   //Byte 3
   //Bit                76543210765432107654321076543210         76543210765432107654321076543210
   IF ((#dWordActCycle AND DW#2#00000011000000000000000000000000) = DW#2#00000010000000000000000000000000) THEN
     #tempCount := #tempCount + 1;
   END_IF;
   //Bit                76543210765432107654321076543210         76543210765432107654321076543210
   IF ((#dWordActCycle AND DW#2#00000110000000000000000000000000) = DW#2#00000100000000000000000000000000) THEN
     #tempCount := #tempCount + 1;
   END_IF;
   //Bit                76543210765432107654321076543210         76543210765432107654321076543210
   IF ((#dWordActCycle AND DW#2#00001100000000000000000000000000) = DW#2#00001000000000000000000000000000) THEN
     #tempCount := #tempCount + 1;
   END_IF;
   //Bit                76543210765432107654321076543210         76543210765432107654321076543210
   IF ((#dWordActCycle AND DW#2#00011000000000000000000000000000) = DW#2#00010000000000000000000000000000) THEN
     #tempCount := #tempCount + 1;
   END_IF;
   //Bit                76543210765432107654321076543210         76543210765432107654321076543210
   IF ((#dWordActCycle AND DW#2#00110000000000000000000000000000) = DW#2#00100000000000000000000000000000) THEN
     #tempCount := #tempCount + 1;
   END_IF;
   //Bit                76543210765432107654321076543210         76543210765432107654321076543210
   IF ((#dWordActCycle AND DW#2#01100000000000000000000000000000) = DW#2#01000000000000000000000000000000) THEN
     #tempCount := #tempCount + 1;
   END_IF;
   //Bit                76543210765432107654321076543210         76543210765432107654321076543210
   IF ((#dWordActCycle AND DW#2#11000000000000000000000000000000) = DW#2#10000000000000000000000000000000) THEN
     #tempCount := #tempCount + 1;
   END_IF;
   //Bit                 76543210765432107654321076543210         76543210765432107654321076543210
   IF (((#dWordActCycle AND DW#2#10000000000000000000000000000000) = DW#2#00000000000000000000000000000000)
     AND ((#statDWordPrevCycle AND DW#2#00000000000000000000000000000001) = DW#2#00000000000000000000000000000001))
   THEN
     #tempCount := #tempCount + 1;
   END_IF;

   // Copy DWord actual cycle to DWord previous cycle
   #statDWordPrevCycle := #dWordActCycle;

   //Output
   #countFalInDWord := #tempCount;
END_FUNCTION_BLOCK

FUNCTION_BLOCK "LGF_CountRisInDWordFB"   // FB10004, SCL
{ S7_Optimized_Access := 'TRUE' }
VERSION : 0.1
   VAR_INPUT
      dWordActCycle : DWord;   // Double word in which the rising edges are counted
   END_VAR
   VAR_OUTPUT
      countRisInDWord : Int;   // Number of rising edges in the double word
   END_VAR
   VAR
      statDWordPrevCycle : DWord;   // Double word from the previous cycle
   END_VAR
   VAR_TEMP
      tempCount : Int;
   END_VAR
BEGIN
   //=============================================================================
   // SIEMENS AG
   // (c)Copyright 2017
   //-----------------------------------------------------------------------------
   // Library:       LGF (Library General Functions)
   // Tested with:   CPU1212C DC/DC/DC FW:V4.2
   // Engineering:   TIA Portal V14 Update 1
   // Restrictions:  -
   // Requirements:  PLC (S7-1200 / S7-1500)
   // Functionality: Detects rising edges in variables of type DWORD
   //-----------------------------------------------------------------------------
   // Change log table:
   // Version  Date        In charge / Changes applied
   // 01.00.00 16.01.2019  Siemens Industry Online Support
   //                      First released version
   //=============================================================================

   // Initialization
   #tempCount := 0;

   //Byte 0
   //Bit                76543210765432107654321076543210         76543210765432107654321076543210
   IF ((#dWordActCycle AND DW#2#00000000000000000000000000000011) = DW#2#00000000000000000000000000000001) THEN
     #tempCount := #tempCount + 1;
   END_IF;
   //Bit                76543210765432107654321076543210         76543210765432107654321076543210
   IF ((#dWordActCycle AND DW#2#00000000000000000000000000000110) = DW#2#00000000000000000000000000000010) THEN
     #tempCount := #tempCount + 1;
   END_IF;
   //Bit                76543210765432107654321076543210         76543210765432107654321076543210
   IF ((#dWordActCycle AND DW#2#00000000000000000000000000001100) = DW#2#00000000000000000000000000000100) THEN
     #tempCount := #tempCount + 1;
   END_IF;
   //Bit                76543210765432107654321076543210         76543210765432107654321076543210
   IF ((#dWordActCycle AND DW#2#00000000000000000000000000011000) = DW#2#00000000000000000000000000001000) THEN
     #tempCount := #tempCount + 1;
   END_IF;
   //Bit                76543210765432107654321076543210         76543210765432107654321076543210
   IF ((#dWordActCycle AND DW#2#00000000000000000000000000110000) = DW#2#00000000000000000000000000010000) THEN
     #tempCount := #tempCount + 1;
   END_IF;
   //Bit                76543210765432107654321076543210         76543210765432107654321076543210
   IF ((#dWordActCycle AND DW#2#00000000000000000000000001100000) = DW#2#00000000000000000000000000100000) THEN
     #tempCount := #tempCount + 1;
   END_IF;
   //Bit                76543210765432107654321076543210         76543210765432107654321076543210
   IF ((#dWordActCycle AND DW#2#00000000000000000000000011000000) = DW#2#00000000000000000000000001000000) THEN
     #tempCount := #tempCount + 1;
   END_IF;
   //Bit                76543210765432107654321076543210         76543210765432107654321076543210
   IF ((#dWordActCycle AND DW#2#00000000000000000000000110000000) = DW#2#00000000000000000000000010000000) THEN
     #tempCount := #tempCount + 1;
   END_IF;

   //Byte 1
   //Bit                76543210765432107654321076543210         76543210765432107654321076543210
   IF ((#dWordActCycle AND DW#2#00000000000000000000001100000000) = DW#2#00000000000000000000000100000000) THEN
     #tempCount := #tempCount + 1;
   END_IF;
   //Bit                76543210765432107654321076543210         76543210765432107654321076543210
   IF ((#dWordActCycle AND DW#2#00000000000000000000011000000000) = DW#2#00000000000000000000001000000000) THEN
     #tempCount := #tempCount + 1;
   END_IF;
   //Bit                76543210765432107654321076543210         76543210765432107654321076543210
   IF ((#dWordActCycle AND DW#2#00000000000000000000110000000000) = DW#2#00000000000000000000010000000000) THEN
     #tempCount := #tempCount + 1;
   END_IF;
   //Bit                76543210765432107654321076543210         76543210765432107654321076543210
   IF ((#dWordActCycle AND DW#2#00000000000000000001100000000000) = DW#2#00000000000000000000100000000000) THEN
     #tempCount := #tempCount + 1;
   END_IF;
   //Bit                76543210765432107654321076543210         76543210765432107654321076543210
   IF ((#dWordActCycle AND DW#2#00000000000000000011000000000000) = DW#2#00000000000000000001000000000000) THEN
     #tempCount := #tempCount + 1;
   END_IF;
   //Bit                76543210765432107654321076543210         76543210765432107654321076543210
   IF ((#dWordActCycle AND DW#2#00000000000000000110000000000000) = DW#2#00000000000000000010000000000000) THEN
     #tempCount := #tempCount + 1;
   END_IF;
   //Bit                76543210765432107654321076543210         76543210765432107654321076543210
   IF ((#dWordActCycle AND DW#2#00000000000000001100000000000000) = DW#2#00000000000000000100000000000000) THEN
     #tempCount := #tempCount + 1;
   END_IF;
   //Bit                76543210765432107654321076543210         76543210765432107654321076543210
   IF ((#dWordActCycle AND DW#2#00000000000000011000000000000000) = DW#2#00000000000000001000000000000000) THEN
     #tempCount := #tempCount + 1;
   END_IF;

   //Byte 2
   //Bit                76543210765432107654321076543210         76543210765432107654321076543210
   IF ((#dWordActCycle AND DW#2#00000000000000110000000000000000) = DW#2#00000000000000010000000000000000) THEN
     #tempCount := #tempCount + 1;
   END_IF;
   //Bit                76543210765432107654321076543210         76543210765432107654321076543210
   IF ((#dWordActCycle AND DW#2#00000000000001100000000000000000) = DW#2#00000000000000100000000000000000) THEN
     #tempCount := #tempCount + 1;
   END_IF;
   //Bit                76543210765432107654321076543210         76543210765432107654321076543210
   IF ((#dWordActCycle AND DW#2#00000000000011000000000000000000) = DW#2#00000000000001000000000000000000) THEN
     #tempCount := #tempCount + 1;
   END_IF;
   //Bit                76543210765432107654321076543210         76543210765432107654321076543210
   IF ((#dWordActCycle AND DW#2#00000000000110000000000000000000) = DW#2#00000000000010000000000000000000) THEN
     #tempCount := #tempCount + 1;
   END_IF;
   //Bit                76543210765432107654321076543210         76543210765432107654321076543210
   IF ((#dWordActCycle AND DW#2#00000000001100000000000000000000) = DW#2#00000000000100000000000000000000) THEN
     #tempCount := #tempCount + 1;
   END_IF;
   //Bit                76543210765432107654321076543210         76543210765432107654321076543210
   IF ((#dWordActCycle AND DW#2#00000000011000000000000000000000) = DW#2#00000000001000000000000000000000) THEN
     #tempCount := #tempCount + 1;
   END_IF;
   //Bit                76543210765432107654321076543210         76543210765432107654321076543210
   IF ((#dWordActCycle AND DW#2#00000000110000000000000000000000) = DW#2#00000000010000000000000000000000) THEN
     #tempCount := #tempCount + 1;
   END_IF;
   //Bit                76543210765432107654321076543210         76543210765432107654321076543210
   IF ((#dWordActCycle AND DW#2#00000001100000000000000000000000) = DW#2#00000000100000000000000000000000) THEN
     #tempCount := #tempCount + 1;
   END_IF;

   //Byte 3
   //Bit                76543210765432107654321076543210         76543210765432107654321076543210
   IF ((#dWordActCycle AND DW#2#00000011000000000000000000000000) = DW#2#00000001000000000000000000000000) THEN
     #tempCount := #tempCount + 1;
   END_IF;
   //Bit                76543210765432107654321076543210         76543210765432107654321076543210
   IF ((#dWordActCycle AND DW#2#00000110000000000000000000000000) = DW#2#00000010000000000000000000000000) THEN
     #tempCount := #tempCount + 1;
   END_IF;
   //Bit                76543210765432107654321076543210         76543210765432107654321076543210
   IF ((#dWordActCycle AND DW#2#00001100000000000000000000000000) = DW#2#00000100000000000000000000000000) THEN
     #tempCount := #tempCount + 1;
   END_IF;
   //Bit                76543210765432107654321076543210         76543210765432107654321076543210
   IF ((#dWordActCycle AND DW#2#00011000000000000000000000000000) = DW#2#00001000000000000000000000000000) THEN
     #tempCount := #tempCount + 1;
   END_IF;
   //Bit                76543210765432107654321076543210         76543210765432107654321076543210
   IF ((#dWordActCycle AND DW#2#00110000000000000000000000000000) = DW#2#00010000000000000000000000000000) THEN
     #tempCount := #tempCount + 1;
   END_IF;
   //Bit                76543210765432107654321076543210         76543210765432107654321076543210
   IF ((#dWordActCycle AND DW#2#01100000000000000000000000000000) = DW#2#00100000000000000000000000000000) THEN
     #tempCount := #tempCount + 1;
   END_IF;
   //Bit                76543210765432107654321076543210         76543210765432107654321076543210
   IF ((#dWordActCycle AND DW#2#11000000000000000000000000000000) = DW#2#01000000000000000000000000000000) THEN
     #tempCount := #tempCount + 1;
   END_IF;
   //Bit                 76543210765432107654321076543210         76543210765432107654321076543210
   IF (((#dWordActCycle AND DW#2#10000000000000000000000000000000) = DW#2#10000000000000000000000000000000)
     AND ((#statDWordPrevCycle AND DW#2#00000000000000000000000000000001) = DW#2#00000000000000000000000000000000))
   THEN
     #tempCount := #tempCount + 1;
   END_IF;

   // Copy DWord actual cycle to DWord previous cycle
   #statDWordPrevCycle := #dWordActCycle;

   //Output
   #countRisInDWord := #tempCount;
END_FUNCTION_BLOCK

// folder: Phisical_functions/LGF/3 Comperator operations

FUNCTION "LGF_CompareVariant" : Bool   // FC10005, SCL
{ S7_Optimized_Access := 'FALSE' }
   VAR_OUTPUT
      error : Bool;
      statusID : UInt;
      status : Word;
   END_VAR
   VAR_IN_OUT
      variable1 : Variant;   // First variable
      variable2 : Variant;   // Second variable
   END_VAR
   VAR_TEMP
      tempVariable1Size : DInt;
      tempVariable2Size : DInt;
      tempCounter : DInt;
      tempVariable1ToBytes : Array[1..#MAX_LENGTH] of Byte;
      tempVariable2ToBytes : Array[1..#MAX_LENGTH] of Byte;
      tempSerializeRet : Int;   // Errorcode. Negative if function fails
   END_VAR
   // Ret_Val : TRUE: equal; FALSE: not equal;
   VAR CONSTANT
      NO_ERROR : Word := 16#0000;
      NO_CURRENT_JOBS : Word := 16#7000;
      ERROR_IN_THIS_BLOCK : UInt := 1;
      ERROR_SERIALIZE : UInt := 2;
      MAX_LENGTH : Int := 200;   // Max. length of PLC datatype in Bytes
   END_VAR
BEGIN
   //=============================================================================
   // SIEMENS AG
   // (c)Copyright 2017
   //-----------------------------------------------------------------------------
   // Library:       LGF (Library General Functions)
   // Tested with:   CPU1212C DC/DC/DC FW:V4.2
   // Engineering:   TIA Portal V14 Update 1
   // Restrictions:  -
   // Requirements:  PLC (S7-1200 / S7-1500)
   // Functionality: Compare the datatypes and values up to a max lengh of 200 Bytes
   //                of the connected variables.
   //                If at least one value of an element is not identical -->
   //                set function result = false
   //-----------------------------------------------------------------------------
   // Change log table:
   // Version Date         In charge / Changes applied
   // 01.00.00 03.09.2015  Siemens Industry Online Support
   //                      First released version
   // 01.00.01 11.02.2015  Siemens Industry Online Support
   //                      Bug fix
   // 01.00.02 02.01.2017  Siemens Industry Online Support
   //                      Upgrade: TIA V14 Update 1
   // 01.00.03 17.08.2018  Siemens Industry Online Support
   //                      Upgrade: TIA V15 Update 2
   // 01.00.04 23.11.2018  Siemens Industry Online Support
   //                      Upgrade: TIA V15.1
   //=============================================================================

   // Set "No current job" #status
   #error := false;
   #statusID := #ERROR_IN_THIS_BLOCK;
   #status := #NO_CURRENT_JOBS;

   // Initialisation of function result
   #LGF_CompareVariant := false;

   // Check if the datatypes of the connected tags are identical
   IF TypeOf(#variable1) = TypeOf(#variable2)
   THEN
     #tempVariable1Size := 0;
     #tempSerializeRet := Serialize(SRC_VARIABLE := #variable1, // convert variable Wert1 to array of byte
                                    DEST_ARRAY => #tempVariable1ToBytes,
                                    POS := #tempVariable1Size);

   // Check return value of SERIALIZE
   IF #tempSerializeRet <> 0
     THEN
       #error := true;
       #statusID := #ERROR_SERIALIZE;
       #status := INT_TO_WORD(#tempSerializeRet);
       RETURN; // Finish function if conversion fails

     ELSE
       #tempVariable2Size := 0;
       // Convert variable Wert2 to array of byte
       #tempSerializeRet := Serialize(SRC_VARIABLE := #variable2,
                                      DEST_ARRAY => #tempVariable2ToBytes,
                                      POS := #tempVariable2Size);

       // Check return value of SERIALIZE
       IF #tempSerializeRet <> 0
       THEN
         #error := true;
         #statusID := #ERROR_SERIALIZE;
         #status := INT_TO_WORD(#tempSerializeRet);
         RETURN; // Finish function if conversion fails
       ELSE

         // Compare size of both variables
         IF #tempVariable1Size = #tempVariable2Size
         THEN
           #tempCounter := 1;

           // Compare values of temp. array elements of bytes
           WHILE #tempCounter <= #tempVariable1Size DO

             // Compare bytes till difference detected
             IF #tempVariable1ToBytes[#tempCounter] = #tempVariable2ToBytes[#tempCounter]    
             THEN
               #tempCounter := #tempCounter + 1; // Or end of array reached
             ELSE
               EXIT;
             END_IF;

           END_WHILE;

           #tempCounter := #tempCounter - 1;
           #LGF_CompareVariant := #tempCounter = #tempVariable1Size; // Assign function result

         END_IF;
       END_IF;
     END_IF;
   END_IF;

   #status := #NO_ERROR;
END_FUNCTION

FUNCTION "LGF_CompareReal" : Bool   // FC10037, SCL
{ S7_Optimized_Access := 'TRUE' }
VERSION : 0.1
   VAR_INPUT
      valueA : Real;   // Number to be compared.
      valueB : Real;   // Number to be compared.
   END_VAR
   VAR_OUTPUT
      error : Bool;   // 0: No error. / 1: Error
      status : Word;   // Error information.
   END_VAR
   // Ret_Val : -
   VAR CONSTANT
      EPSILON : Real := 1.0E-06;   // Accuracy with which the two numbers are considered equal
      MAX_RANGE_REAL : Real := 3.402823E+38;   // Maximum range of a REAL number
      ERROR_OVERFLOW : Word := 16#8601;   // Maximum range of a REAL number exceeded
      NO_ERROR : Word := 16#0000;   // No error.
   END_VAR
BEGIN
   //=============================================================================
   // Siemens AG
   // (c)Copyright 2017
   //-----------------------------------------------------------------------------
   // Library:       LGF (Library General Functions)
   // Tested with:   CPU1212C DC/DC/DC FW:V4.2
   // Engineering:   TIA Portal V14 Upd 1
   // Restrictions:  -
   // Requirements:  PLC (S7-1200 / S7-1500)
   // Functionality: This function checks real numbers for parity
   //-----------------------------------------------------------------------------
   // Change log table:
   // Version  Date        In charge / Changes applied
   // 01.00.00 13.01.2017  Siemens Industry Online Support
   //                      First released version
   // 01.00.01 17.08.2018  Siemens Industry Online Support
   //                      Upgrade: TIA V15 Update 2
   // 01.00.02 23.11.2018  Siemens Industry Online Support
   //                      Upgrade: TIA V15.1
   //-----------------------------------------------------------------------------
   //Status Codes: 16#0000 - no error
   //              16#8601 - |valueA|+|valueB| exceeds the maximum range of REAL
   //=============================================================================

   // Reset outputs
   #error := FALSE;
   #status := #NO_ERROR;

   // Initialisation of function result
   #LGF_CompareReal := FALSE;

   // Check |valueA|+|valueB| does not exceed the maximum range of REAL
   IF (ABS(#valueA) + ABS(#valueB)) > #MAX_RANGE_REAL THEN
       #error := TRUE;
       #status := #ERROR_OVERFLOW;
       RETURN;
   END_IF;

   // Approximation
   #LGF_CompareReal := ABS(#valueA - #valueB) <= (#EPSILON * (ABS(#valueA) + ABS(#valueB)));
END_FUNCTION

// folder: Phisical_functions/LGF/4 Math operations

FUNCTION_BLOCK "LGF_MinMaxHistory"   // FB10012, SCL
{ S7_Optimized_Access := 'TRUE' }
   VAR_INPUT
      variable : LReal;
      reset : Bool;
   END_VAR
   VAR_OUTPUT
      minValue : LReal := 1.7976931348623157e+308;
      maxValue : LReal := -1.7976931348623157e+308;
   END_VAR
   VAR
      statMinValue : LReal := 1.7976931348623157e+308;
      statMaxValue : LReal := -1.7976931348623157e+308;
   END_VAR
   VAR CONSTANT
      LREAL_MAX : LReal := 1.7976931348623157e+308;
      LREAL_MIN : LReal := -1.7976931348623157e+308;
   END_VAR
BEGIN
   //=============================================================================
   // SIEMENS AG
   // (c)Copyright 2017
   //-----------------------------------------------------------------------------
   // Library:       LGF (Library General Functions)
   // Tested with:   CPU1212C DC/DC/DC FW:V4.2
   // Engineering:   TIA Portal V14 Update 1
   // Restrictions:  -
   // Requirements:  PLC (S7-1200 / S7-1500)
   // Functionality: This function block saves the minimum and maximum value,
   //                since the start of the block.
   //-----------------------------------------------------------------------------
   // Change log table:
   // Version  Date        In charge / Changes applied
   // 01.00.00 19.08.2015  Siemens Industry Online Support
   //                      First released version
   // 01.00.01 02.01.2017  Siemens Industry Online Support
   //                      Upgrade: TIA Portal V14 Update 1
   //                      Code optimization
   // 01.00.02 17.08.2018  Siemens Industry Online Support
   //                      Upgrade: TIA V15 Update 2
   // 01.00.03 23.11.2018  Siemens Industry Online Support
   //                      Upgrade: TIA V15.1
   //=============================================================================

   // Save min value
   IF (#variable < #statMinValue) THEN
     #statMinValue := #variable;
   END_IF;

   // Save max value
   IF (#variable > #statMaxValue ) THEN
     #statMaxValue := #variable;
   END_IF;

   // If reset is TRUE, min and max value are set to 0
   IF (#reset = TRUE)  THEN
     #statMinValue := #LREAL_MAX;
     #statMaxValue := #LREAL_MIN;
   ELSE
     ;
   END_IF;

   // Ouptput of min and max value
   #minValue := #statMinValue;
   #maxValue := #statMaxValue;
END_FUNCTION_BLOCK

FUNCTION_BLOCK "LGF_Integration"   // FB10043, SCL
{ S7_Optimized_Access := 'TRUE' }
VERSION : 0.1
   VAR_INPUT
      value : Real;   // -
      enable : Bool;   // -
      reset : Bool;   // -
   END_VAR
   VAR_OUTPUT
      integral : Real;   // -
      error : Bool;   // -
      statusID : UInt;   // -
      status : Word;   // Status information / -
   END_VAR
   VAR
      statSysTime : DTL;   // -
      statLastTime : DTL;   // -
      statOldValue : Real;   // -
      statIntegral : Real;   // -
      tempValue : Real;   // -
      tempDeltaTimeT : Time;   // -
      tempDeltaTimeDInt : DInt;   // -
      tempDeltaTimeReal : Real;   // -
      tempRetval : Int;   // -
   END_VAR
   VAR CONSTANT
      ZERO : Real := 0.0;
      NO_ERROR : Word := 16#0000;   // -
      NO_CURRENT_JOBS : Word := 16#7000;   // -
      ERROR_IN_THIS_BLOCK : UInt := 1;   // error in this block
      ERROR_RD_SYS_T : UInt := 2;   // error in RD_SYS_T
   END_VAR
BEGIN
   //=============================================================================
   // SIEMENS AG
   // (c)Copyright 2017
   //-----------------------------------------------------------------------------
   // Library:       LGF (Library General Functions)
   // Tested with:   CPU1212C DC/DC/DC FW:V4.2
   // Engineering:   TIA Portal V14 Upd 1
   // Restrictions:  -
   // Requirements:  PLC (S7-1200 / S7-1500)
   // Functionality: The input value will be integrated.
   //                
   //-----------------------------------------------------------------------------
   // Change log table:
   // Version  Date        In charge Changes applied
   // 01.00.00 17.02.2017  Siemens Industry Online Support
   //                      First released version
   // 01.00.01 17.08.2018  Siemens Industry Online Support
   //                      Upgrade: TIA V15 Update 2
   // 01.00.02 23.11.2018  Siemens Industry Online Support
   //                      Upgrade: TIA V15.1
   //-----------------------------------------------------------------------------
   //=============================================================================

   // Initialization
   #error := FALSE;
   #statusID := #NO_ERROR;
   #status := #NO_CURRENT_JOBS;

   // Reset 
   IF #reset = true THEN
     #integral := #ZERO;
     #statOldValue := #ZERO;
     #statIntegral := #ZERO;
     RETURN;
   END_IF;

   // Write input value to temp variable
   #tempValue := #value;

   // Read system time
   #tempRetval := RD_SYS_T(OUT => #statSysTime);

   // Error Handling read system time
   IF (#tempRetval > 1) THEN
     #error := TRUE;
     #statusID := #ERROR_RD_SYS_T;
     #status := INT_TO_WORD(#tempRetval);
     RETURN;
   END_IF;

   // Calculate time difference between last and actual time
   #tempDeltaTimeT := #statSysTime - #statLastTime;

   // Convert times difference to REAL
   #tempDeltaTimeDInt := TIME_TO_DINT(#tempDeltaTimeT);
   #tempDeltaTimeReal := DINT_TO_REAL(#tempDeltaTimeDInt);

   // Convert in seconds
   #tempDeltaTimeReal := #tempDeltaTimeReal / 1000.0;

   // Write actual to last time
   #statLastTime := #statSysTime;

   IF NOT #enable = true THEN
     #statOldValue := #ZERO;
     RETURN;
   END_IF;

   // Add LastScalIn to ScalIn
   #tempValue := #tempValue + #statOldValue;

   // Save last input
   #statOldValue := #value;

   // Divide in half statScalIn
   #tempValue := #tempValue / 2.0;

   // Multiply with Delta Time
   #tempValue := #tempValue * #tempDeltaTimeReal;

   // Calculate new integral
   #statIntegral := #statIntegral + #tempValue;

   // Write outputs
   #integral := #statIntegral;
   #status := #NO_ERROR;
END_FUNCTION_BLOCK

FUNCTION "LGF_RandomInt" : Int   // FC2, SCL
{ S7_Optimized_Access := 'TRUE' }
   VAR_INPUT
      minValue : Int;   // minimal Value random can reach
      maxValue : Int;   // maximal Value random can reach
   END_VAR
   VAR_OUTPUT
      error : Bool;
      statusID : UInt;
      status : Word;
   END_VAR
   VAR_TEMP
      tempTime : DTL;
      tempTimeStatus : Int;
      tempRandomValue : Int;
      tempNormReal : Real;
   END_VAR
   VAR CONSTANT
      NO_ERROR : Word := 16#0000;
      NO_CURRENT_JOBS : Word := 16#7000;
      MAX_LESS_MIN : Word := 16#8200;
      ERROR_IN_THIS_BLOCK : UInt := 1;
      ERROR_RD_SYS_T : UInt := 2;
      MIN_INT : DInt := -32768;
      MAX_INT : DInt := 32767;
   END_VAR
BEGIN
   //=============================================================================
   // Siemens AG
   // (c)Copyright 2017
   //-----------------------------------------------------------------------------
   // Library:       LGF (Library General Functions)
   // Tested with:   CPU1212C DC/DC/DC FW:V4.2
   // Engineering:   TIA Portal V13 SP1 Upd 4
   // Restrictions:  -
   // Requirements:  PLC (S7-1200 / S7-1500)
   // Functionality: This function generates random numbers in defined limits
   //                (Datatype Int)
   //-----------------------------------------------------------------------------
   // Change log table:
   // Version  Date        In charge / Changes applied
   // 01.00.00 19.08.2015  Siemens Industry Online Support
   //                      First released version
   // 01.00.01 02.01.2017  Siemens Industry Online Support
   //                      Upgrade: TIA Portal V14 Update 1
   // 01.00.02 17.08.2018  Siemens Industry Online Support
   //                      Upgrade: TIA V15 Update 2
   // 01.00.03 23.11.2018  Siemens Industry Online Support
   //                      Upgrade: TIA V15.1
   //-----------------------------------------------------------------------------
   //Status Codes:
   // 16#7000:  No current jobs
   // 16#0000:  Job finished; Note: There is no "Busy"-Status because the block
   //           is finished within a single cycle
   // 16#8200:  maxValue is samller then minValue 
   //=============================================================================

   //Set "No current job" status
   #error := false;
   #statusID := #ERROR_IN_THIS_BLOCK;
   #status := #NO_CURRENT_JOBS;

   //Check if the maximal Value is less than the minimal value
   IF (#minValue > #maxValue) THEN
     #error := true;
     #statusID := #ERROR_IN_THIS_BLOCK;
     #status := #MAX_LESS_MIN;
     #LGF_RandomInt := 0;
     RETURN;
   END_IF;

   //Read system time
   #tempTimeStatus := RD_SYS_T(#tempTime);

   IF (#tempTimeStatus <> 0) THEN
     #error := true;
     #statusID := #ERROR_RD_SYS_T;
     #status := INT_TO_WORD(#tempTimeStatus);
     #LGF_RandomInt := 0;
     RETURN;
   END_IF;

   //Callculate a random-start-value depending on the time
   #tempRandomValue.%B1 := #tempTime.NANOSECOND.%B0;
   #tempRandomValue.%B0 := #tempTime.NANOSECOND.%B1;

   //adapt the calculated random number to the given number span
   #tempNormReal := NORM_X(MIN := #MIN_INT, VALUE := #tempRandomValue, MAX := #MAX_INT);
   #LGF_RandomInt := SCALE_X(MIN := #minValue, VALUE := #tempNormReal, MAX := #maxValue);

   #status := #NO_ERROR;
END_FUNCTION

FUNCTION "LGF_Factorial" : DInt   // FC9, SCL
{ S7_Optimized_Access := 'TRUE' }
VERSION : 0.1
   VAR_INPUT
      n : Int;   // Natural number
   END_VAR
   VAR_OUTPUT
      status : Word;   // Status
      error : Bool;   // Error
   END_VAR
   VAR_TEMP
      tempFactorial : DInt;   // Temp Factorial
      tempIndex : Int;   // Temp index
   END_VAR
   // Ret_Val : Calculated factorial
   VAR CONSTANT
      NO_ERROR : Word := 16#0000;   // Status no error
      NO_CURRENT_JOBS : Word := 16#7000;   // Status no current jobs
      WRONG_VALUE_RANGE : Word := 16#8101;   // Status wrong value range for input value
   END_VAR
BEGIN
   //=============================================================================
   // Siemens AG
   // (c)Copyright 2017
   //-----------------------------------------------------------------------------
   // Library:       LGF (Library General Functions)
   // Tested with:   CPU1212C DC/DC/DC FW:V4.2
   // Engineering:   TIA Portal V14 SP1 Upd 5
   // Restrictions:  -
   // Requirements:  PLC (S7-1200 / S7-1500)
   // Functionality: This program calculates factorial values from 1 to 12.
   //-----------------------------------------------------------------------------
   // Change log table:
   // Version  Date        In charge / Changes applied
   // 01.00.00 03.07.2018  Siemens Industry Online Support
   //                      First released version
   // 01.00.01 17.08.2018  Siemens Industry Online Support
   //                      Upgrade: TIA V15 Update 2
   // 01.00.02 23.11.2018  Siemens Industry Online Support
   //                      Upgrade: TIA V15.1
   //-----------------------------------------------------------------------------
   //Status Codes:
   // 16#0000:  Job finished   // Note: There is no "Busy"-Status because the
   //           block is finished within a single cycle
   // 16#8101:  Outside value range ( factorial until 12 is possible)
   //=============================================================================

   #error := FALSE;
   #status := #NO_CURRENT_JOBS;

   IF (#n < 13)
     AND (#n >= 0)
   THEN
     IF (#n = 0)
     THEN
       #tempFactorial := 1;
     ELSE
       #tempFactorial := 1;
       FOR #tempIndex := 1 TO #n DO
         #tempFactorial := #tempFactorial * #tempIndex;
       END_FOR;
     END_IF;

     #error := FALSE; // No errors
     #status := #NO_ERROR;

   ELSE
     #tempFactorial := 0;
     #error := TRUE;
     #status := #WRONG_VALUE_RANGE;
   END_IF;

   #LGF_Factorial := #tempFactorial;
END_FUNCTION

FUNCTION "LGF_MatrixAddition" : Void   // FC10007, SCL
{ S7_Optimized_Access := 'TRUE' }
   VAR_INPUT
      matrix1 : Array[*, *] of Real;   // first summand
      matrix2 : Array[*, *] of Real;   // second summand
   END_VAR
   VAR_OUTPUT
      matrixResult : Array[*, *] of Real;   // result matrix
      error : Bool;
      statusID : UInt;
      status : Word;
   END_VAR
   VAR_TEMP
      tempMatrix1LowerBound1Dim : DInt;   // -
      tempMatrix1LowerBound2Dim : DInt;   // -
      tempMatrix1UpperBound1Dim : DInt;   // -
      tempMatrix1UpperBound2Dim : DInt;   // -
      tempMatrix2LowerBound1Dim : DInt;   // -
      tempMatrix2LowerBound2Dim : DInt;   // -
      tempMatrix2UpperBound1Dim : DInt;   // -
      tempMatrix2UpperBound2Dim : DInt;   // -
      tempResultMatrixLowerBound1Dim : DInt;   // -
      tempResultMatrixLowerBound2Dim : DInt;   // -
      tempResultMatrixUpperBound1Dim : DInt;   // -
      tempResultMatrixUpperBound2Dim : DInt;   // -
      tempCounterDim1 : Int;   // -
      tempCounterDim2 : Int;   // -
   END_VAR
   VAR CONSTANT
      NO_ERROR : Word := 16#0000;   // No errors.
      ERROR_LOWER_BOUND_NOT_EQUAL : Word := 16#8200;   // Lower bounds of matrices are not equal.
      ERROR_UPPER_BOUND_NOT_EQUAL : Word := 16#8201;   // Upper bounds of matrices are not equal.
      ERROR_IN_THIS_BLOCK : UInt := 1;   // statusID: Error in this block.
   END_VAR
BEGIN
   //=============================================================================
   // SIEMENS AG
   // (c)Copyright 2017
   //-----------------------------------------------------------------------------
   // Library:       LGF (Library General Functions)
   // Tested with:   CPU1212C DC/DC/DC FW:V4.2
   // Engineering:   TIA Portal V14 Update 1
   // Restrictions:  -
   // Requirements:  PLC (S7-1200 / S7-1500)
   // Functionality: This function add up matrices.
   //-----------------------------------------------------------------------------
   // Change log table:
   // Version  Date        In charge / Changes applied
   // 01.00.00 19.08.2015  Siemens Industry Online Support
   //                      First released version
   // 01.00.01 02.01.2017  Siemens Industry Online Support
   //                      Upgrade: TIA Portal V14 Update 1
   // 02.00.00 06.02.2017  Siemens Industry Online Support
   //                      Functionality using Array[*,*]
   // 02.00.01 17.08.2018  Siemens Industry Online Support
   //                      Upgrade: TIA V15 Update 2
   // 02.00.02 23.11.2018  Siemens Industry Online Support
   //                      Upgrade: TIA V15.1
   //=============================================================================

   //Set "No error" status
   #error := false;
   #statusID := #ERROR_IN_THIS_BLOCK;
   #status := #NO_ERROR;

   // Init resultMatrix
   #matrixResult[0, 0] := 0.0;

   //Determine the size of the matrices
   // Lower bound dimension 1
   #tempMatrix1LowerBound1Dim := LOWER_BOUND(ARR := #matrix1, DIM := 1);
   #tempMatrix2LowerBound1Dim := LOWER_BOUND(ARR := #matrix2, DIM := 1);
   #tempResultMatrixLowerBound1Dim := LOWER_BOUND(ARR := #matrixResult, DIM := 1);
   // Lower bound dimension 2
   #tempMatrix1LowerBound2Dim := LOWER_BOUND(ARR := #matrix1, DIM := 2);
   #tempMatrix2LowerBound2Dim := LOWER_BOUND(ARR := #matrix2, DIM := 2);
   #tempResultMatrixLowerBound2Dim := LOWER_BOUND(ARR := #matrixResult, DIM := 2);
   // Upper bound dimension 1
   #tempMatrix1UpperBound1Dim := UPPER_BOUND(ARR := #matrix1, DIM := 1);
   #tempMatrix2UpperBound1Dim := UPPER_BOUND(ARR := #matrix2, DIM := 1);
   #tempResultMatrixUpperBound1Dim := UPPER_BOUND(ARR := #matrixResult, DIM := 1);
   // Upper bound dimension 2
   #tempMatrix1UpperBound2Dim := UPPER_BOUND(ARR := #matrix1, DIM := 2);
   #tempMatrix2UpperBound2Dim := UPPER_BOUND(ARR := #matrix2, DIM := 2);
   #tempResultMatrixUpperBound2Dim := UPPER_BOUND(ARR := #matrixResult, DIM := 2);

   // Check the lower bound of all matrices
   IF (#tempMatrix1LowerBound1Dim <> #tempMatrix2LowerBound1Dim) OR (#tempMatrix1LowerBound1Dim <> #tempResultMatrixLowerBound1Dim) OR
     (#tempMatrix1LowerBound2Dim <> #tempMatrix2LowerBound2Dim) OR (#tempMatrix1LowerBound2Dim <> #tempResultMatrixLowerBound2Dim) THEN
     #error := TRUE;
     #status := #ERROR_LOWER_BOUND_NOT_EQUAL;
     RETURN;
   END_IF;
   // Check the upper bound of all matrices
   IF (#tempMatrix1UpperBound1Dim <> #tempMatrix2UpperBound1Dim) OR (#tempMatrix1UpperBound1Dim <> #tempResultMatrixUpperBound1Dim) OR
     (#tempMatrix1UpperBound2Dim <> #tempMatrix2UpperBound2Dim) OR (#tempMatrix1UpperBound2Dim <> #tempResultMatrixUpperBound2Dim) THEN
     #error := TRUE;
     #status := #ERROR_UPPER_BOUND_NOT_EQUAL;
     RETURN;
   END_IF;

   // Addition of two matrices
   FOR #tempCounterDim1 := #tempMatrix1LowerBound1Dim TO #tempMatrix1UpperBound1Dim DO
     FOR #tempCounterDim2 := #tempMatrix1LowerBound2Dim TO #tempMatrix1UpperBound2Dim DO
       #matrixResult[#tempCounterDim1, #tempCounterDim2] := #matrix1[#tempCounterDim1, #tempCounterDim2] + #matrix2[#tempCounterDim1, #tempCounterDim2];
     END_FOR;
   END_FOR;
END_FUNCTION

FUNCTION "LGF_MatrixInverse" : Void   // FC10008, SCL
{ S7_Optimized_Access := 'TRUE' }
   VAR_INPUT
      matrix : Array[*, *] of Real;   // input matrix
   END_VAR
   VAR_OUTPUT
      matrixResult : Array[*, *] of Real;   // output matrix
      error : Bool;
      statusID : UInt;
      status : Word;
   END_VAR
   VAR_TEMP
      tempCounterDim2 : Int;   // -
      tempCounterDim1 : Int;   // -
      tempMatrixLowerBound1Dim : DInt;   // -
      tempMatrixLowerBound2Dim : DInt;   // -
      tempMatrixUpperBound1Dim : DInt;   // -
      tempMatrixUpperBound2Dim : DInt;   // -
      tempResultMatrixLowerBound1Dim : DInt;   // -
      tempResultMatrixLowerBound2Dim : DInt;   // -
      tempResultMatrixUpperBound1Dim : DInt;   // -
      tempResultMatrixUpperBound2Dim : DInt;   // -
      tempColumns : DInt;   // -
      tempRows : DInt;   // -
      tempK : DInt;   // -
      tempI : DInt;   // -
      tempJ : DInt;   // -
   END_VAR
   VAR CONSTANT
      NO_ERROR : Word := 16#0000;   // No error.
      ERROR_LOWER_BOUND_NOT_EQUAL : Word := 16#8200;   // Lower bounds of matrices are not equal.
      ERROR_UPPER_BOUND_NOT_EQUAL : Word := 16#8201;   // Upper bounds of matrices are not equal.
      ERROR_NOT_SQUARE_MATRIX : Word := 16#8202;   // Input matrix is not a square matrix.
      ERROR_ALGORITHM_NOT_POSSIBLE : Word := 16#8203;   // Algorithm not possible for the input matrix.
      ERROR_IN_THIS_BLOCK : UInt := 1;   // statusID: error in this block.
   END_VAR
BEGIN
   //=============================================================================
   // SIEMENS AG
   // (c)Copyright 2017
   //-----------------------------------------------------------------------------
   // Library:       LGF (Library General Functions)
   // Tested with:   CPU1212C DC/DC/DC FW:V4.2
   // Engineering:   TIA Portal V14 Update 1
   // Restrictions:  -
   // Requirements:  PLC (S7-1200 / S7-1500)
   // Functionality: This function inverses matrices. Inversion of regulary,
   //                quadratic Matrix with the Shipley-Coleman method.
   //-----------------------------------------------------------------------------
   // Change log table:
   // Version  Date        In charge / Changes applied
   // 01.00.00 19.08.2015  Siemens Industry Online Support
   //                      First released version
   // 01.00.01 02.01.2017  Siemens Industry Online Support
   //                      Upgrade: TIA Portal V14 Update 1
   // 02.00.00 06.02.2017  Siemens Industry Online Support
   //                      Functionality using Array[*,*]
   // 02.00.01 17.08.2018  Siemens Industry Online Support
   //                      Upgrade: TIA V15 Update 2
   // 02.00.02 23.11.2018  Siemens Industry Online Support
   //                      Upgrade: TIA V15.1
   //=============================================================================

   //Set "No error" status
   #error := false;
   #statusID := #ERROR_IN_THIS_BLOCK;
   #status := #NO_ERROR;

   // Initialize result matrix
   #matrixResult[0, 0] := 0.0;

   //Determine the size of the matrices
   // Lower bound dimension 1
   #tempMatrixLowerBound1Dim := LOWER_BOUND(ARR := #matrix, DIM := 1);
   #tempResultMatrixLowerBound1Dim := LOWER_BOUND(ARR := #matrixResult, DIM := 1);
   // Lower bound dimension 2
   #tempMatrixLowerBound2Dim := LOWER_BOUND(ARR := #matrix, DIM := 2);
   #tempResultMatrixLowerBound2Dim := LOWER_BOUND(ARR := #matrixResult, DIM := 2);
   // Upper bound dimension 1
   #tempMatrixUpperBound1Dim := UPPER_BOUND(ARR := #matrix, DIM := 1);
   #tempResultMatrixUpperBound1Dim := UPPER_BOUND(ARR := #matrixResult, DIM := 1);
   // Upper bound dimension 2
   #tempMatrixUpperBound2Dim := UPPER_BOUND(ARR := #matrix, DIM := 2);
   #tempResultMatrixUpperBound2Dim := UPPER_BOUND(ARR := #matrixResult, DIM := 2);

   // Count the columns of input matrix
   IF #tempMatrixLowerBound2Dim = 0 THEN
     #tempColumns := #tempMatrixUpperBound2Dim + 1;
   ELSE
     #tempColumns := (#tempMatrixUpperBound2Dim - #tempMatrixLowerBound2Dim) + 1;
   END_IF;
   // Count the rows of input matrix
   IF #tempMatrixLowerBound1Dim = 0 THEN
     #tempRows := #tempMatrixUpperBound1Dim + 1;
   ELSE
     #tempRows := (#tempMatrixUpperBound1Dim - #tempMatrixLowerBound1Dim) + 1;
   END_IF;
   // Check whether input matrix is a square matrix
   IF #tempRows <> #tempColumns THEN
     #error := TRUE;
     #status := #ERROR_NOT_SQUARE_MATRIX;
     RETURN;
   END_IF;

   // Output matrix must have same lower bounds as the input matrix. (Same array size)
   IF (#tempMatrixLowerBound1Dim <> #tempResultMatrixLowerBound1Dim) OR (#tempMatrixLowerBound2Dim <> #tempResultMatrixLowerBound2Dim) THEN
     #error := TRUE;
     #status := #ERROR_LOWER_BOUND_NOT_EQUAL;
     RETURN;
   END_IF;
   // Output matrix must have same upper bounds as the input matrix. (Same array size)
   IF (#tempMatrixUpperBound1Dim <> #tempResultMatrixUpperBound1Dim) OR (#tempMatrixUpperBound2Dim <> #tempResultMatrixUpperBound2Dim) THEN
     #error := TRUE;
     #status := #ERROR_UPPER_BOUND_NOT_EQUAL;
     RETURN;
   END_IF;

   // Negate the input matrix and copy to output matrix.
   FOR #tempCounterDim1 := #tempMatrixLowerBound1Dim TO #tempMatrixUpperBound1Dim DO
     FOR #tempCounterDim2 := #tempMatrixLowerBound2Dim TO #tempMatrixUpperBound2Dim DO
       #matrixResult[#tempCounterDim1, #tempCounterDim2] := - #matrix[#tempCounterDim1, #tempCounterDim2];
     END_FOR;
   END_FOR;

   //Outside loop - relegation of "Main" diagonal
   FOR #tempK := #tempMatrixLowerBound2Dim TO #tempMatrixUpperBound2Dim DO

     // Avoid a division by zero --> Error: Algorithm does not work for the input matrix.
     IF #matrixResult[#tempK, #tempK] = 0.0 THEN
       #error := TRUE;
       #status := #ERROR_ALGORITHM_NOT_POSSIBLE;
       RETURN;
     ELSE
       //Calculation of Pivot-element.
       #matrixResult[#tempK, #tempK] :=
       (-1 / #matrixResult[#tempK, #tempK]);
     END_IF;

     //Calculation of elemente in the Pivot-column.
     FOR #tempI := #tempMatrixLowerBound2Dim TO #tempMatrixUpperBound2Dim DO
       IF #tempI <> #tempK THEN
         #matrixResult[#tempI, #tempK] :=
         #matrixResult[#tempI, #tempK] * #matrixResult[#tempK, #tempK];
       END_IF;
     END_FOR;

     // Convert-calculation of elements, which are NOT in the Pivot-rolumn AND NOT in the Pivot-row.
     FOR #tempI := #tempMatrixLowerBound1Dim TO #tempMatrixUpperBound1Dim DO

       IF #tempI <> #tempK THEN
         FOR #tempJ := #tempMatrixLowerBound2Dim TO #tempMatrixUpperBound2Dim DO
           IF #tempJ <> #tempK THEN
             #matrixResult[#tempI, #tempJ] :=
             #matrixResult[#tempI, #tempJ] + #matrixResult[#tempI, #tempK] * #matrixResult[#tempK, #tempJ];
           END_IF;
         END_FOR;
       END_IF;
     END_FOR;

     //Calculation of elements in the Pivot-row.
     FOR #tempJ := #tempMatrixLowerBound2Dim TO #tempMatrixUpperBound2Dim DO
       IF #tempJ <> #tempK THEN
         #matrixResult[#tempK, #tempJ] :=
         #matrixResult[#tempK, #tempJ] * #matrixResult[#tempK, #tempK];
       END_IF;
     END_FOR;
   END_FOR;
END_FUNCTION

FUNCTION "LGF_MatrixMultiplication" : Void   // FC10009, SCL
{ S7_Optimized_Access := 'TRUE' }
   VAR_INPUT
      matrix1 : Array[*, *] of Real;   // First matrix.
      matrix2 : Array[*, *] of Real;   // Second matrix.
   END_VAR
   VAR_OUTPUT
      matrixResult : Array[*, *] of Real;   // Output matrix.
      error : Bool;
      statusID : UInt;
      status : Word;
   END_VAR
   VAR_TEMP
      tempMatrix1LowerBound1Dim : DInt;   // -
      tempMatrix1LowerBound2Dim : DInt;   // -
      tempMatrix1UpperBound1Dim : DInt;   // -
      tempMatrix1UpperBound2Dim : DInt;   // -
      tempMatrix2LowerBound1Dim : DInt;   // -
      tempMatrix2LowerBound2Dim : DInt;   // -
      tempMatrix2UpperBound1Dim : DInt;   // -
      tempMatrix2UpperBound2Dim : DInt;   // -
      tempResultMatrixLowerBound1Dim : DInt;   // -
      tempResultMatrixLowerBound2Dim : DInt;   // -
      tempResultMatrixUpperBound1Dim : DInt;   // -
      tempResultMatrixUpperBound2Dim : DInt;   // -
      tempCounterJ : Int;   // -
      tempCounterK : Int;   // -
      tempCounterL : Int;   // -
      tempResult : Real;   // -
   END_VAR
   VAR CONSTANT
      NO_ERROR : Word := 16#0000;   // No error.
      ERROR_WRONG_INPUT_MATRIX : Word := 16#8200;   // Dimension 2 of matrix 1 <> Dimension 1 of matrix 2
      ERROR_WRONG_OUTPUT_MATRIX : Word := 16#8201;   // Dimension 1 <> dimension 1 of matrix 1; Dimension 2 <> dimension 2 of matrix2
      ERROR_IN_THIS_BLOCK : UInt := 1;   // statusID: error in this block.
   END_VAR
BEGIN
   //=============================================================================
   // SIEMENS AG
   // (c)Copyright 2017
   //-----------------------------------------------------------------------------
   // Library:       LGF (Library General Functions)
   // Tested with:   CPU1212C DC/DC/DC FW:V4.2
   // Engineering:   TIA Portal V14 Update 1
   // Restrictions:  -
   // Requirements:  PLC (S7-1200 / S7-1500)
   // Functionality: This function multiplicates matrices.
   //-----------------------------------------------------------------------------
   // Change log table:
   // Version  Date        In charge / Changes applied
   // 01.00.00 19.08.2015  Siemens Industry Online Support
   //                      First released version
   // 01.00.01 02.01.2017  Siemens Industry Online Support
   //                      Upgrade: TIA Portal V14 Update 1
   // 02.00.00 06.02.2017  Siemens Industry Online Support
   //                      Functionality using Array[*,*]
   // 02.00.01 17.08.2018  Siemens Industry Online Support
   //                      Upgrade: TIA V15 Update 2
   // 02.00.02 23.11.2018  Siemens Industry Online Support
   //                      Upgrade: TIA V15.1
   //=============================================================================

   //Set "No error" status
   #error := false;
   #statusID := #ERROR_IN_THIS_BLOCK;
   #status := #NO_ERROR;

   // Initialize the output matrix
   #matrixResult[0, 0] := 0.0;

   //Determine the size of the matrices
   // Lower bound dimension 1
   #tempMatrix1LowerBound1Dim := LOWER_BOUND(ARR := #matrix1, DIM := 1);
   #tempMatrix2LowerBound1Dim := LOWER_BOUND(ARR := #matrix2, DIM := 1);
   #tempResultMatrixLowerBound1Dim := LOWER_BOUND(ARR := #matrixResult, DIM := 1);
   // Lower bound dimension 2
   #tempMatrix1LowerBound2Dim := LOWER_BOUND(ARR := #matrix1, DIM := 2);
   #tempMatrix2LowerBound2Dim := LOWER_BOUND(ARR := #matrix2, DIM := 2);
   #tempResultMatrixLowerBound2Dim := LOWER_BOUND(ARR := #matrixResult, DIM := 2);
   // Upper bound dimension 1
   #tempMatrix1UpperBound1Dim := UPPER_BOUND(ARR := #matrix1, DIM := 1);
   #tempMatrix2UpperBound1Dim := UPPER_BOUND(ARR := #matrix2, DIM := 1);
   #tempResultMatrixUpperBound1Dim := UPPER_BOUND(ARR := #matrixResult, DIM := 1);
   // Upper bound dimension 2
   #tempMatrix1UpperBound2Dim := UPPER_BOUND(ARR := #matrix1, DIM := 2);
   #tempMatrix2UpperBound2Dim := UPPER_BOUND(ARR := #matrix2, DIM := 2);
   #tempResultMatrixUpperBound2Dim := UPPER_BOUND(ARR := #matrixResult, DIM := 2);

   // Matrix one must have the same count of rows as matrix two has columns. Else the multiplication is not possible.
   IF (#tempMatrix1LowerBound2Dim <> #tempMatrix2LowerBound1Dim) OR (#tempMatrix1UpperBound2Dim <> #tempMatrix2UpperBound1Dim) THEN
     #error := true;
     #statusID := #ERROR_IN_THIS_BLOCK;
     #status := #ERROR_WRONG_INPUT_MATRIX;
     RETURN;
   END_IF;
   // Result matrix must have the same number of rows as matrix 1 and the same number of columns as the matrix 2 (same lower and upper bound)
   IF (#tempMatrix1LowerBound1Dim <> #tempResultMatrixLowerBound1Dim) OR (#tempMatrix1UpperBound1Dim <> #tempResultMatrixUpperBound1Dim)
     OR (#tempMatrix2LowerBound2Dim <> #tempResultMatrixLowerBound2Dim) OR (#tempMatrix2UpperBound2Dim <> #tempResultMatrixUpperBound2Dim) THEN
     #error := true;
     #statusID := #ERROR_IN_THIS_BLOCK;
     #status := #ERROR_WRONG_OUTPUT_MATRIX;
     RETURN;
   END_IF;

   // Multiplication
   FOR #tempCounterJ := #tempMatrix1LowerBound1Dim TO #tempMatrix1UpperBound1Dim DO
     FOR #tempCounterK := #tempMatrix2LowerBound2Dim TO #tempMatrix2UpperBound2Dim DO
       #tempResult := 0.0;
       FOR #tempCounterL := #tempMatrix1LowerBound2Dim TO #tempMatrix1UpperBound2Dim DO
         #tempResult := #tempResult + #matrix1[#tempCounterJ, #tempCounterL] * #matrix2[#tempCounterL, #tempCounterK];
       END_FOR;
       #matrixResult[#tempCounterJ, #tempCounterK] := #tempResult;
     END_FOR;
   END_FOR;
END_FUNCTION
